Flt - Depress Man Weld To Continue FB2[301].22'; 9655 '~S001R16CN.I.Wc2SGunFlt - Weld Controller 2 Servo Gun Fault FB2[301].23'; 9656 '~S001R16CN.I.Wc2SGunMtrTempFlt - Cntrl 2 Servo Gun Motor Over Temp FB2[301].24'; 9657 '~S001R16CN.I.Td2MtrFlt - Tip Dress 2 Motor Fault FB2[301].25'; 9658 '~S001R16CN.I.WC2XfmrTempFlt - Weld Cntrl 2 Transformer Over Temp FB2[301].26'; 9659 '~S001R16CN.I.AutoTipChng2Flt - Auto Tip Changer 2 Fault FB2[301].27'; 9660 '~S001R16CN.I.Slr2NotReady - Seal Controller 2 Not Ready FB2[301].28'; 9661 '~S001R16CN.I.Slr2MajorFlt - Seal Controller 2 Major Fault FB2[301].29'; 9662 '~S001R16CN.I.Slr2VolNotOk - Seal Controller 2 Volume Not Ok Fault FB2[301].30'; 9663 '~S001R16CN.I.Slr2PurgeFlt - Seal Controller 2 Purge Fault FB2[301].31'; 9664 '~S001R16CN.I.Slr2DoserNot Filled - Seal Cntrl 2 Doser Not Filled FB2[302].0'; 9665 '~S001R16CN.I.Slr2No2ClnMxr - Seal Cntrl2 No 2C In Mixer Fault FB2[302].1'; 9666 '~S001R16CN.I.Slr2NzlBroken - Seal Controller 2 Nozzle Broken Fault FB2[302].2'; 9667 '~S001R16CN.I.Slr2NozzleChgReq - Seal Cntrl2 Nozzle Change Reqd FB2[302].3'; 9668 '~S001R16CN.I.Slr2CycleInterrupted - Seal Cntrl2 Cycle Interrupted FB2[302].4'; 9669 '~S001R16CN.I.Stdw2Flt - Stud Weld 2 Weld Fault FB2[302].5'; 9670 '~S001R16CN.I.Stdw2DlyExcdd - Stud Weld 2 Time Delay Exceeded Flt FB2[302].6'; 9671 '~S001R16CN.I.Stdw2Maint Reqd - Stud Weld 2 Maintenance Required FB2[302].7'; 9672 '~S001R16CN.I.Stdw2Reject - Stud Weld 2 art Reject Fault FB2[302].8'; 9673 '~S001R16CN.I.Rvt2Flt - Rivet Controller 2 Fault FB2[302].9'; 9674 '~S001R16CN.I.Rvt2DlyExcdd - Rivet Cntrl 2 Time Delay Exceeded Flt FB2[302].10'; 9675 '~S001R16CN.I.AutoPulledTipByp2 - Auto Pulled Tip Bypass 2 FB2[302].11'; 9676 '~S001R16CN.I.StdWld2EquipmentFlt - Stud Weld 2 Equipment Fault FB2[302].12'; 9677 '~S001R16CN.I.StdWld2BrcktNotPresent - Stud Weld 2 Bracket Not Pres FB2[302].13'; 9678 '~S001R16CN.Ix.LsrWldMntrFlt - Seam Geometry/Laser Weld Monitor Flt FB2[302].14'; 9679 '~S001R16CN.Ix.LsrHeadFlt - Laser Head Fault FB2[302].15'; 9680 '~S001R16CN.Ix.LsrGlsFlt - Glass Fault FB2[302].16'; 9681 '~S001R16CN.Ix.LsrWhlFlt - Pressure Wheel Not In Range Fault FB2[302].17'; 9682 '~S001R16CN.Ix.LsrGeoFlt - Seam Geometry/Laser Bad Process Geo Flt FB2[302].18'; 9683 '~S001R16CN.Ix.LsrHdCollFlt - Laser Head Collision Fault FB2[302].19'; 9684 '~S001R16CN.Ix.LsrHdSysFlt - Laser Head System Fault FB2[302].20'; 9685 '~S001R16CN.Ix.LsrHdFar - Laser Head Far Fault FB2[302].21'; 9686 '~S001R16CN.Ix.LsrHdSftCollFlt - Laser Head Software Collision Flt FB2[302].22'; 9687 '~S001R16CN.I.O.TipChngReqd2 - Weld Cntrl 2 Tip Change Required FB2[302].23'; 9688 '~S001R16CN.I.M.NutDetectFlt2 - Nut Welder 2 Nut Detection Fault FB2[302].24'; 9689 '~S001R16CN.I.M.NutProjFlt2 - Nut Welder 2 Weld Not In Tolerance FB2[302].25'; 9690 '~S001R16CN.I.TCWrongToolInStand - Tool Changer Wrong Tool In Stand FB2[302].26'; 9691 '~Spare FB2[302].27'; 9692 '~Spare FB2[302].28'; 9693 '~Spare FB2[302].29'; 9694 '~Spare FB2[302].30'; 9695 '~Spare FB2[302].31'; 9696 '~S001R16CN.I.VisionCommOK - Vision System Comm Fault FB2[303].0'; 9697 '~S001R16CN.I.OutOfTolerance - Vision System Out Of Tolerance FB2[303].1'; 9698 '~S001R16CN.I.MeasureReject - Vision System Measure Reject FB2[303].2'; 9699 '~S001R16CN.I.VisionSysCalibrationFlt - Vision System Calibration Flt FB2[303].3'; 9700 '~S001R16CN.I.VisionSysFlt - Vision System Flt FB2[303].4'; 9701 '~Spare FB2[303].5'; 9702 '~Spare FB2[303].6'; 9703 '~Spare FB2[303].7'; 9704 '~Spare FB2[303].8'; 9705 '~Spare FB2[303].9'; 9706 '~Spare FB2[303].10'; 9707 '~Spare FB2[303].11'; 9708 '~Spare FB2[303].12'; 9709 '~Spare FB2[303].13'; 9710 '~Spare FB2[303].14'; 9711 '~Spare FB2[303].15'; 9712 '~Spare FB2[303].16'; 9713 '~Spare FB2[303].17'; 9714 '~S001R16CN.M.InteruptCyc - Laser Cyc Interupt Cut Wire And Reject Car FB2[303].18'; 9715 '~S001R16CN.M.SuspectPart Inspect Vehicle And Accept Or Reject FB2[303].19'; 9716 '~S001R16 Power Meter High Power Fault Detected FB2[303].20'; 9717 '~S001R16 Power Meter Low Power Fault Detected FB2[303].21'; 9718 '~Spare FB2[303].22'; 9719 '~Spare FB2[303].23'; 9720 '~Spare FB2[303].24'; 9721 '~Spare FB2[303].25'; 9722 '~Spare FB2[303].26'; 9723 '~Spare FB2[303].27'; 9724 '~Spare FB2[303].28'; 9725 '~Spare FB2[303].29'; 9726 '~Spare FB2[303].30'; 9727 '~Spare FB2[303].31'; 9728 '~Spare FB2[304].0'; 9729 '~Spare FB2[304].1'; 9730 '~Spare FB2[304].2'; 9731 '~Spare FB2[304].3'; 9732 '~Spare FB2[304].4'; 9733 '~Spare FB2[304].5'; 9734 '~Spare FB2[304].6'; 9735 '~Spare FB2[304].7'; 9736 '~Spare FB2[304].8'; 9737 '~Spare FB2[304].9'; 9738 '~Spare FB2[304].10'; 9739 '~Spare FB2[304].11'; 9740 '~Spare FB2[304].12'; 9741 '~Spare FB2[304].13'; 9742 '~Spare FB2[304].14'; 9743 '~Spare FB2[304].15'; 9744 '~Spare FB2[304].16'; 9745 '~Spare FB2[304].17'; 9746 '~Spare FB2[304].18'; 9747 '~Spare FB2[304].19'; 9748 '~Spare FB2[304].20'; 9749 '~Spare FB2[304].21'; 9750 '~Spare FB2[304].22'; 9751 '~Spare FB2[304].23'; 9752 '~Spare FB2[304].24'; 9753 '~Spare FB2[304].25'; 9754 '~Spare FB2[304].26'; 9755 '~Spare FB2[304].27'; 9756 '~Spare FB2[304].28'; 9757 '~Spare FB2[304].29'; 9758 '~Spare FB2[304].30'; 9759 '~Spare FB2[304].31'; 9760 '~Spare FB2[305].0'; 9761 '~Spare FB2[305].1'; 9762 '~Spare FB2[305].2'; 9763 '~Spare FB2[305].3'; 9764 '~Spare FB2[305].4'; 9765 '~Spare FB2[305].5'; 9766 '~Spare FB2[305].6'; 9767 '~Spare FB2[305].7'; 9768 '~Spare FB2[305].8'; 9769 '~Spare FB2[305].9'; 9770 '~Spare FB2[305].10'; 9771 '~Spare FB2[305].11'; 9772 '~Spare FB2[305].12'; 9773 '~Spare FB2[305].13'; 9774 '~Spare FB2[305].14'; 9775 '~Spare FB2[305].15'; 9776 '~Spare FB2[305].16'; 9777 '~Spare FB2[305].17'; 9778 '~Spare FB2[305].18'; 9779 '~Spare FB2[305].19'; 9780 '~Spare FB2[305].20'; 9781 '~Spare FB2[305].21'; 9782 '~Spare FB2[305].22'; 9783 '~Spare FB2[305].23'; 9784 '~Spare FB2[305].24'; 9785 '~Spare FB2[305].25'; 9786 '~Spare FB2[305].26'; 9787 '~Spare FB2[305].27'; 9788 '~Spare FB2[305].28'; 9789 '~Spare FB2[305].29'; 9790 '~Spare FB2[305].30'; 9791 '~Spare FB2[305].31'; 9792 '~Spare FB2[306].0'; 9793 '~Spare FB2[306].1'; 9794 '~Spare FB2[306].2'; 9795 '~Spare FB2[306].3'; 9796 '~Spare FB2[306].4'; 9797 '~Spare FB2[306].5'; 9798 '~Spare FB2[306].6'; 9799 '~Spare FB2[306].7'; 9800 '~Spare FB2[306].8'; 9801 '~Spare FB2[306].9'; 9802 '~Spare FB2[306].10'; 9803 '~Spare FB2[306].11'; 9804 '~Spare FB2[306].12'; 9805 '~Spare FB2[306].13'; 9806 '~Spare FB2[306].14'; 9807 '~Spare FB2[306].15'; 9808 '~Spare FB2[306].16'; 9809 '~Spare FB2[306].17'; 9810 '~Spare FB2[306].18'; 9811 '~Spare FB2[306].19'; 9812 '~Spare FB2[306].20'; 9813 '~Spare FB2[306].21'; 9814 '~Spare FB2[306].22'; 9815 '~Spare FB2[306].23'; 9816 '~Spare FB2[306].24'; 9817 '~Spare FB2[306].25'; 9818 '~Spare FB2[306].26'; 9819 '~Spare FB2[306].27'; 9820 '~Spare FB2[306].28'; 9821 '~Spare FB2[306].29'; 9822 '~Spare FB2[306].30'; 9823 '~Spare FB2[306].31'; 9824 '~Spare FB2[307].0'; 9825 '~Spare FB2[307].1'; 9826 '~Spare FB2[307].2'; 9827 '~Spare FB2[307].3'; 9828 '~Spare FB2[307].4'; 9829 '~Spare FB2[307].5'; 9830 '~Spare FB2[307].6'; 9831 '~Spare FB2[307].7'; 9832 '~Spare FB2[307].8'; 9833 '~Spare FB2[307].9'; 9834 '~Spare FB2[307].10'; 9835 '~Spare FB2[307].11'; 9836 '~Spare FB2[307].12'; 9837 '~Spare FB2[307].13'; 9838 '~Spare FB2[307].14'; 9839 '~Spare FB2[307].15'; 9840 '~Spare FB2[307].16'; 9841 '~Spare FB2[307].17'; 9842 '~Spare FB2[307].18'; 9843 '~Spare FB2[307].19'; 9844 '~Spare FB2[307].20'; 9845 '~Spare FB2[307].21'; 9846 '~Spare FB2[307].22'; 9847 '~Spare FB2[307].23'; 9848 '~Spare FB2[307].24'; 9849 '~Spare FB2[307].25'; 9850 '~Spare FB2[307].26'; 9851 '~Spare FB2[307].27'; 9852 '~Spare FB2[307].28'; 9853 '~Spare FB2[307].29'; 9854 '~Spare FB2[307].30'; 9855 '~Spare FB2[307].31'; 9856 '~Spare FB2[308].0'; 9857 '~Spare FB2[308].1'; 9858 '~Spare FB2[308].2'; 9859 '~Spare FB2[308].3'; 9860 '~Spare FB2[308].4'; 9861 '~Spare FB2[308].5'; 9862 '~Spare FB2[308].6'; 9863 '~Spare FB2[308].7'; 9864 '~Spare FB2[308].8'; 9865 '~Spare FB2[308].9'; 9866 '~Spare FB2[308].10'; 9867 '~Spare FB2[308].11'; 9868 '~Spare FB2[308].12'; 9869 '~Spare FB2[308].13'; 9870 '~Spare FB2[308].14'; 9871 '~Spare FB2[308].15'; 9872 '~Spare FB2[308].16'; 9873 '~Spare FB2[308].17'; 9874 '~Spare FB2[308].18'; 9875 '~Spare FB2[308].19'; 9876 '~Spare FB2[308].20'; 9877 '~Spare FB2[308].21'; 9878 '~Spare FB2[308].22'; 9879 '~Spare FB2[308].23'; 9880 '~Spare FB2[308].24'; 9881 '~Spare FB2[308].25'; 9882 '~Spare FB2[308].26'; 9883 '~Spare FB2[308].27'; 9884 '~Spare FB2[308].28'; 9885 '~Spare FB2[308].29'; 9886 '~Spare FB2[308].30'; 9887 '~Spare FB2[308].31'; 9888 '~Spare FB2[309].0'; 9889 '~Spare FB2[309].1'; 9890 '~Spare FB2[309].2'; 9891 '~Spare FB2[309].3'; 9892 '~Spare FB2[309].4'; 9893 '~Spare FB2[309].5'; 9894 '~Spare FB2[309].6'; 9895 '~Spare FB2[309].7'; 9896 '~Spare FB2[309].8'; 9897 '~Spare FB2[309].9'; 9898 '~Spare FB2[309].10'; 9899 '~Spare FB2[309].11'; 9900 '~Spare FB2[309].12'; 9901 '~Spare FB2[309].13'; 9902 '~Spare FB2[309].14'; 9903 '~Spare FB2[309].15'; 9904 '~Spare FB2[309].16'; 9905 '~Spare FB2[309].17'; 9906 '~Spare FB2[309].18'; 9907 '~Spare FB2[309].19'; 9908 '~Spare FB2[309].20'; 9909 '~Spare FB2[309].21'; 9910 '~Spare FB2[309].22'; 9911 '~Spare FB2[309].23'; 9912 '~Spare FB2[309].24'; 9913 '~Spare FB2[309].25'; 9914 '~Spare FB2[309].26'; 9915 '~Spare FB2[309].27'; 9916 '~Spare FB2[309].28'; 9917 '~Spare FB2[309].29'; 9918 '~Spare FB2[309].30'; 9919 '~Spare FB2[309].31'; 9920 '~Spare FB2[310].0'; 9921 '~Spare FB2[310].1'; 9922 '~Spare FB2[310].2'; 9923 '~Spare FB2[310].3'; 9924 '~Spare FB2[310].4'; 9925 '~Spare FB2[310].5'; 9926 '~Spare FB2[310].6'; 9927 '~Spare FB2[310].7'; 9928 '~Spare FB2[310].8'; 9929 '~Spare FB2[310].9'; 9930 '~Spare FB2[310].10'; 9931 '~Spare FB2[310].11'; 9932 '~Spare FB2[310].12'; 9933 '~Spare FB2[310].13'; 9934 '~Spare FB2[310].14'; 9935 '~Spare FB2[310].15'; 9936 '~Spare FB2[310].16'; 9937 '~Spare FB2[310].17'; 9938 '~Spare FB2[310].18'; 9939 '~Spare FB2[310].19'; 9940 '~Spare FB2[310].20'; 9941 '~Spare FB2[310].21'; 9942 '~Spare FB2[310].22'; 9943 '~Spare FB2[310].23'; 9944 '~Spare FB2[310].24'; 9945 '~Spare FB2[310].25'; 9946 '~Spare FB2[310].26'; 9947 '~Spare FB2[310].27'; 9948 '~Spare FB2[310].28'; 9949 '~Spare FB2[310].29'; 9950 '~Spare FB2[310].30'; 9951 '~Spare FB2[310].31'; 9952 '~Spare FB2[311].0'; 9953 '~Spare FB2[311].1'; 9954 '~Spare FB2[311].2'; 9955 '~Spare FB2[311].3'; 9956 '~Spare FB2[311].4'; 9957 '~Spare FB2[311].5'; 9958 '~Spare FB2[311].6'; 9959 '~Spare FB2[311].7'; 9960 '~Spare FB2[311].8'; 9961 '~Spare FB2[311].9'; 9962 '~Spare FB2[311].10'; 9963 '~Spare FB2[311].11'; 9964 '~Spare FB2[311].12'; 9965 '~Spare FB2[311].13'; 9966 '~Spare FB2[311].14'; 9967 '~Spare FB2[311].15'; 9968 '~Spare FB2[311].16'; 9969 '~Spare FB2[311].17'; 9970 '~Spare FB2[311].18'; 9971 '~Spare FB2[311].19'; 9972 '~Spare FB2[311].20'; 9973 '~Spare FB2[311].21'; 9974 '~Spare FB2[311].22'; 9975 '~Spare FB2[311].23'; 9976 '~Spare FB2[311].24'; 9977 '~Spare FB2[311].25'; 9978 '~Spare FB2[311].26'; 9979 '~Spare FB2[311].27'; 9980 '~Spare FB2[311].28'; 9981 '~Spare FB2[311].29'; 9982 '~Spare FB2[311].30'; 9983 '~Spare FB2[311].31'; 9984 '~Spare FB2[312].0'; 9985 '~Spare FB2[312].1'; 9986 '~Spare FB2[312].2'; 9987 '~Spare FB2[312].3'; 9988 '~Spare FB2[312].4'; 9989 '~Spare FB2[312].5'; 9990 '~Spare FB2[312].6'; 9991 '~Spare FB2[312].7'; 9992 '~Spare FB2[312].8'; 9993 '~Spare FB2[312].9'; 9994 '~Spare FB2[312].10'; 9995 '~Spare FB2[312].11'; 9996 '~Spare FB2[312].12'; 9997 '~Spare FB2[312].13'; 9998 '~Spare FB2[312].14'; 9999 '~Spare FB2[312].15'; 10000 '**Local Message Display**'

